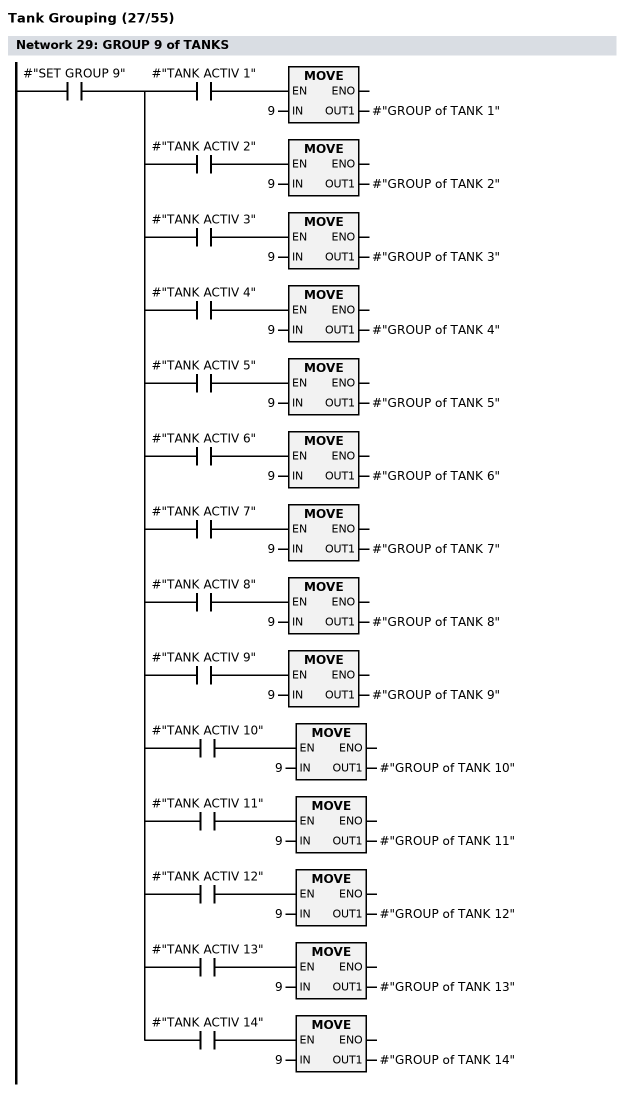
   RUNG wire#powerrail
      Contact( #"SET GROUP 9" )
      wire#w1
      Contact( #"TANK ACTIV 1" )
      Move(in := 9, out1 => #"GROUP of TANK 1")
   END_RUNG
   RUNG wire#w1
      Contact( #"TANK ACTIV 2" )
      Move(in := 9, out1 => #"GROUP of TANK 2")
   END_RUNG
   RUNG wire#w1
      Contact( #"TANK ACTIV 3" )
      Move(in := 9, out1 => #"GROUP of TANK 3")
   END_RUNG
   RUNG wire#w1
      Contact( #"TANK ACTIV 4" )
      Move(in := 9, out1 => #"GROUP of TANK 4")
   END_RUNG
   RUNG wire#w1
      Contact( #"TANK ACTIV 5" )
      Move(in := 9, out1 => #"GROUP of TANK 5")
   END_RUNG
   RUNG wire#w1
      Contact( #"TANK ACTIV 6" )
      Move(in := 9, out1 => #"GROUP of TANK 6")
   END_RUNG
   RUNG wire#w1
      Contact( #"TANK ACTIV 7" )
      Move(in := 9, out1 => #"GROUP of TANK 7")
   END_RUNG
   RUNG wire#w1
      Contact( #"TANK ACTIV 8" )
      Move(in := 9, out1 => #"GROUP of TANK 8")
   END_RUNG
   RUNG wire#w1
      Contact( #"TANK ACTIV 9" )
      Move(in := 9, out1 => #"GROUP of TANK 9")
   END_RUNG
   RUNG wire#w1
      Contact( #"TANK ACTIV 10" )
      Move(in := 9, out1 => #"GROUP of TANK 10")
   END_RUNG
   RUNG wire#w1
      Contact( #"TANK ACTIV 11" )
      Move(in := 9, out1 => #"GROUP of TANK 11")
   END_RUNG
   RUNG wire#w1
      Contact( #"TANK ACTIV 12" )
      Move(in := 9, out1 => #"GROUP of TANK 12")
   END_RUNG
   RUNG wire#w1
      Contact( #"TANK ACTIV 13" )
      Move(in := 9, out1 => #"GROUP of TANK 13")
   END_RUNG
   RUNG wire#w1
      Contact( #"TANK ACTIV 14" )
      Move(in := 9, out1 => #"GROUP of TANK 14")
   END_RUNG
   // the same network as SCL:
   IF #"SET GROUP 9" AND #"TANK ACTIV 1" THEN #"GROUP of TANK 1" := 9; END_IF;
   IF #"SET GROUP 9" AND #"TANK ACTIV 2" THEN #"GROUP of TANK 2" := 9; END_IF;
   IF #"SET GROUP 9" AND #"TANK ACTIV 3" THEN #"GROUP of TANK 3" := 9; END_IF;
   IF #"SET GROUP 9" AND #"TANK ACTIV 4" THEN #"GROUP of TANK 4" := 9; END_IF;
   IF #"SET GROUP 9" AND #"TANK ACTIV 5" THEN #"GROUP of TANK 5" := 9; END_IF;
   IF #"SET GROUP 9" AND #"TANK ACTIV 6" THEN #"GROUP of TANK 6" := 9; END_IF;
   IF #"SET GROUP 9" AND #"TANK ACTIV 7" THEN #"GROUP of TANK 7" := 9; END_IF;
   IF #"SET GROUP 9" AND #"TANK ACTIV 8" THEN #"GROUP of TANK 8" := 9; END_IF;
   IF #"SET GROUP 9" AND #"TANK ACTIV 9" THEN #"GROUP of TANK 9" := 9; END_IF;
   IF #"SET GROUP 9" AND #"TANK ACTIV 10" THEN #"GROUP of TANK 10" := 9; END_IF;
   IF #"SET GROUP 9" AND #"TANK ACTIV 11" THEN #"GROUP of TANK 11" := 9; END_IF;
   IF #"SET GROUP 9" AND #"TANK ACTIV 12" THEN #"GROUP of TANK 12" := 9; END_IF;
   IF #"SET GROUP 9" AND #"TANK ACTIV 13" THEN #"GROUP of TANK 13" := 9; END_IF;
   IF #"SET GROUP 9" AND #"TANK ACTIV 14" THEN #"GROUP of TANK 14" := 9; END_IF;
END_REGION

REGION Network 30: GROUP 10 of TANKS
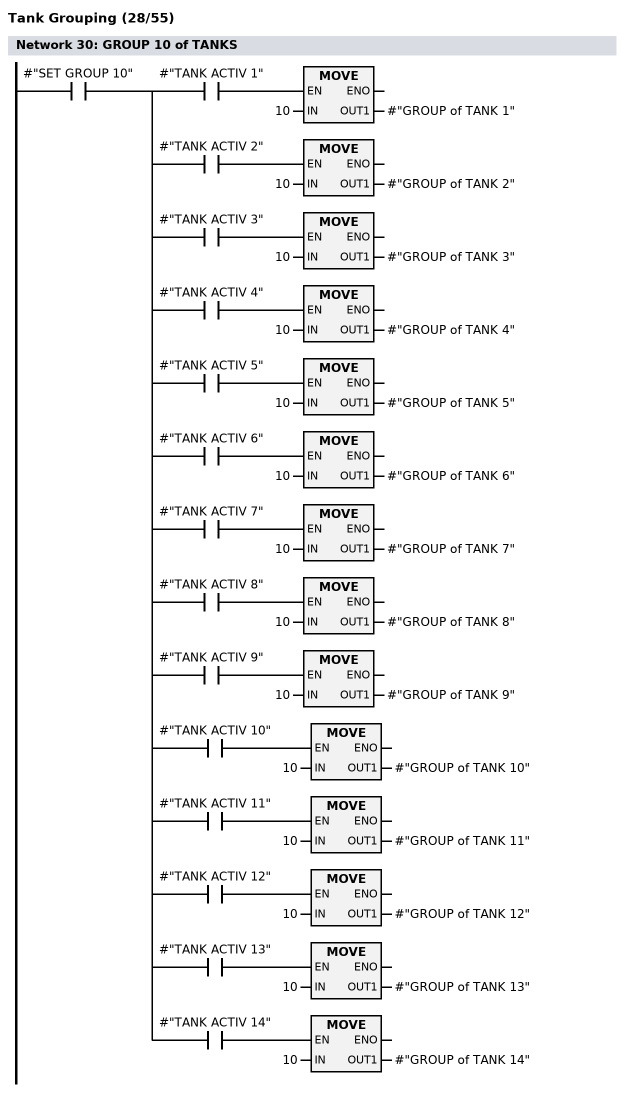
   RUNG wire#powerrail
      Contact( #"SET GROUP 10" )
      wire#w1
      Contact( #"TANK ACTIV 1" )
      Move(in := 10, out1 => #"GROUP of TANK 1")
   END_RUNG
   RUNG wire#w1
      Contact( #"TANK ACTIV 2" )
      Move(in := 10, out1 => #"GROUP of TANK 2")
   END_RUNG
   RUNG wire#w1
      Contact( #"TANK ACTIV 3" )
      Move(in := 10, out1 => #"GROUP of TANK 3")
   END_RUNG
   RUNG wire#w1
      Contact( #"TANK ACTIV 4" )
      Move(in := 10, out1 => #"GROUP of TANK 4")
   END_RUNG
   RUNG wire#w1
      Contact( #"TANK ACTIV 5" )
      Move(in := 10, out1 => #"GROUP of TANK 5")
   END_RUNG
   RUNG wire#w1
      Contact( #"TANK ACTIV 6" )
      Move(in := 10, out1 => #"GROUP of TANK 6")
   END_RUNG
   RUNG wire#w1
      Contact( #"TANK ACTIV 7" )
      Move(in := 10, out1 => #"GROUP of TANK 7")
   END_RUNG
   RUNG wire#w1
      Contact( #"TANK ACTIV 8" )
      Move(in := 10, out1 => #"GROUP of TANK 8")
   END_RUNG
   RUNG wire#w1
      Contact( #"TANK ACTIV 9" )
      Move(in := 10, out1 => #"GROUP of TANK 9")
   END_RUNG
   RUNG wire#w1
      Contact( #"TANK ACTIV 10" )
      Move(in := 10, out1 => #"GROUP of TANK 10")
   END_RUNG
   RUNG wire#w1
      Contact( #"TANK ACTIV 11" )
      Move(in := 10, out1 => #"GROUP of TANK 11")
   END_RUNG
   RUNG wire#w1
      Contact( #"TANK ACTIV 12" )
      Move(in := 10, out1 => #"GROUP of TANK 12")
   END_RUNG
   RUNG wire#w1
      Contact( #"TANK ACTIV 13" )
      Move(in := 10, out1 => #"GROUP of TANK 13")
   END_RUNG
   RUNG wire#w1
      Contact( #"TANK ACTIV 14" )
      Move(in := 10, out1 => #"GROUP of TANK 14")
   END_RUNG
   // the same network as SCL:
   IF #"SET GROUP 10" AND #"TANK ACTIV 1" THEN #"GROUP of TANK 1" := 10; END_IF;
   IF #"SET GROUP 10" AND #"TANK ACTIV 2" THEN #"GROUP of TANK 2" := 10; END_IF;
   IF #"SET GROUP 10" AND #"TANK ACTIV 3" THEN #"GROUP of TANK 3" := 10; END_IF;
   IF #"SET GROUP 10" AND #"TANK ACTIV 4" THEN #"GROUP of TANK 4" := 10; END_IF;
   IF #"SET GROUP 10" AND #"TANK ACTIV 5" THEN #"GROUP of TANK 5" := 10; END_IF;
   IF #"SET GROUP 10" AND #"TANK ACTIV 6" THEN #"GROUP of TANK 6" := 10; END_IF;
   IF #"SET GROUP 10" AND #"TANK ACTIV 7" THEN #"GROUP of TANK 7" := 10; END_IF;
   IF #"SET GROUP 10" AND #"TANK ACTIV 8" THEN #"GROUP of TANK 8" := 10; END_IF;
   IF #"SET GROUP 10" AND #"TANK ACTIV 9" THEN #"GROUP of TANK 9" := 10; END_IF;
   IF #"SET GROUP 10" AND #"TANK ACTIV 10" THEN #"GROUP of TANK 10" := 10; END_IF;
   IF #"SET GROUP 10" AND #"TANK ACTIV 11" THEN #"GROUP of TANK 11" := 10; END_IF;
   IF #"SET GROUP 10" AND #"TANK ACTIV 12" THEN #"GROUP of TANK 12" := 10; END_IF;
   IF #"SET GROUP 10" AND #"TANK ACTIV 13" THEN #"GROUP of TANK 13" := 10; END_IF;
   IF #"SET GROUP 10" AND #"TANK ACTIV 14" THEN #"GROUP of TANK 14" := 10; END_IF;
END_REGION

REGION Network 31: GROUP 11 of TANKS
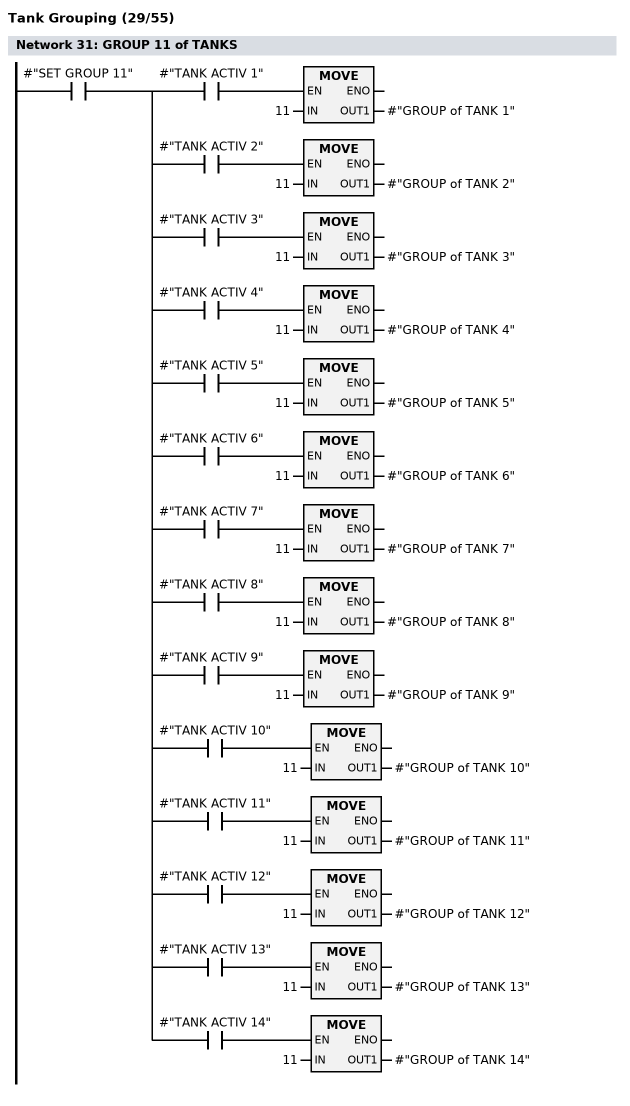
   RUNG wire#powerrail
      Contact( #"SET GROUP 11" )
      wire#w1
      Contact( #"TANK ACTIV 1" )
      Move(in := 11, out1 => #"GROUP of TANK 1")
   END_RUNG
   RUNG wire#w1
      Contact( #"TANK ACTIV 2" )
      Move(in := 11, out1 => #"GROUP of TANK 2")
   END_RUNG
   RUNG wire#w1
      Contact( #"TANK ACTIV 3" )
      Move(in := 11, out1 => #"GROUP of TANK 3")
   END_RUNG
   RUNG wire#w1
      Contact( #"TANK ACTIV 4" )
      Move(in := 11, out1 => #"GROUP of TANK 4")
   END_RUNG
   RUNG wire#w1
      Contact( #"TANK ACTIV 5" )
      Move(in := 11, out1 => #"GROUP of TANK 5")
   END_RUNG
   RUNG wire#w1
      Contact( #"TANK ACTIV 6" )
      Move(in := 11, out1 => #"GROUP of TANK 6")
   END_RUNG
   RUNG wire#w1
      Contact( #"TANK ACTIV 7" )
      Move(in := 11, out1 => #"GROUP of TANK 7")
   END_RUNG
   RUNG wire#w1
      Contact( #"TANK ACTIV 8" )
      Move(in := 11, out1 => #"GROUP of TANK 8")
   END_RUNG
   RUNG wire#w1
      Contact( #"TANK ACTIV 9" )
      Move(in := 11, out1 => #"GROUP of TANK 9")
   END_RUNG
   RUNG wire#w1
      Contact( #"TANK ACTIV 10" )
      Move(in := 11, out1 => #"GROUP of TANK 10")
   END_RUNG
   RUNG wire#w1
      Contact( #"TANK ACTIV 11" )
      Move(in := 11, out1 => #"GROUP of TANK 11")
   END_RUNG
   RUNG wire#w1
      Contact( #"TANK ACTIV 12" )
      Move(in := 11, out1 => #"GROUP of TANK 12")
   END_RUNG
   RUNG wire#w1
      Contact( #"TANK ACTIV 13" )
      Move(in := 11, out1 => #"GROUP of TANK 13")
   END_RUNG
   RUNG wire#w1
      Contact( #"TANK ACTIV 14" )
      Move(in := 11, out1 => #"GROUP of TANK 14")
   END_RUNG
   // the same network as SCL:
   IF #"SET GROUP 11" AND #"TANK ACTIV 1" THEN #"GROUP of TANK 1" := 11; END_IF;
   IF #"SET GROUP 11" AND #"TANK ACTIV 2" THEN #"GROUP of TANK 2" := 11; END_IF;
   IF #"SET GROUP 11" AND #"TANK ACTIV 3" THEN #"GROUP of TANK 3" := 11; END_IF;
   IF #"SET GROUP 11" AND #"TANK ACTIV 4" THEN #"GROUP of TANK 4" := 11; END_IF;
   IF #"SET GROUP 11" AND #"TANK ACTIV 5" THEN #"GROUP of TANK 5" := 11; END_IF;
   IF #"SET GROUP 11" AND #"TANK ACTIV 6" THEN #"GROUP of TANK 6" := 11; END_IF;
   IF #"SET GROUP 11" AND #"TANK ACTIV 7" THEN #"GROUP of TANK 7" := 11; END_IF;
   IF #"SET GROUP 11" AND #"TANK ACTIV 8" THEN #"GROUP of TANK 8" := 11; END_IF;
   IF #"SET GROUP 11" AND #"TANK ACTIV 9" THEN #"GROUP of TANK 9" := 11; END_IF;
   IF #"SET GROUP 11" AND #"TANK ACTIV 10" THEN #"GROUP of TANK 10" := 11; END_IF;
   IF #"SET GROUP 11" AND #"TANK ACTIV 11" THEN #"GROUP of TANK 11" := 11; END_IF;
   IF #"SET GROUP 11" AND #"TANK ACTIV 12" THEN #"GROUP of TANK 12" := 11; END_IF;
   IF #"SET GROUP 11" AND #"TANK ACTIV 13" THEN #"GROUP of TANK 13" := 11; END_IF;
   IF #"SET GROUP 11" AND #"TANK ACTIV 14" THEN #"GROUP of TANK 14" := 11; END_IF;
END_REGION

REGION Network 32: GROUP 12 of TANKS
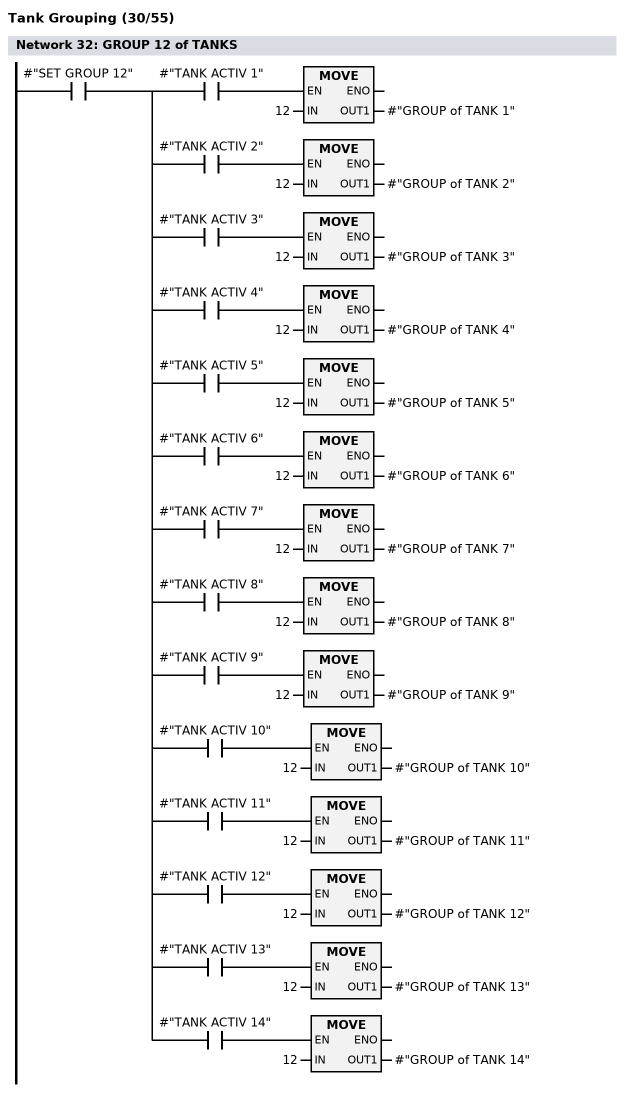
   RUNG wire#powerrail
      Contact( #"SET GROUP 12" )
      wire#w1
      Contact( #"TANK ACTIV 1" )
      Move(in := 12, out1 => #"GROUP of TANK 1")
   END_RUNG
   RUNG wire#w1
      Contact( #"TANK ACTIV 2" )
      Move(in := 12, out1 => #"GROUP of TANK 2")
   END_RUNG
   RUNG wire#w1
      Contact( #"TANK ACTIV 3" )
      Move(in := 12, out1 => #"GROUP of TANK 3")
   END_RUNG
   RUNG wire#w1
      Contact( #"TANK ACTIV 4" )
      Move(in := 12, out1 => #"GROUP of TANK 4")
   END_RUNG
   RUNG wire#w1
      Contact( #"TANK ACTIV 5" )
      Move(in := 12, out1 => #"GROUP of TANK 5")
   END_RUNG
   RUNG wire#w1
      Contact( #"TANK ACTIV 6" )
      Move(in := 12, out1 => #"GROUP of TANK 6")
   END_RUNG
   RUNG wire#w1
      Contact( #"TANK ACTIV 7" )
      Move(in := 12, out1 => #"GROUP of TANK 7")
   END_RUNG
   RUNG wire#w1
      Contact( #"TANK ACTIV 8" )
      Move(in := 12, out1 => #"GROUP of TANK 8")
   END_RUNG
   RUNG wire#w1
      Contact( #"TANK ACTIV 9" )
      Move(in := 12, out1 => #"GROUP of TANK 9")
   END_RUNG
   RUNG wire#w1
      Contact( #"TANK ACTIV 10" )
      Move(in := 12, out1 => #"GROUP of TANK 10")
   END_RUNG
   RUNG wire#w1
      Contact( #"TANK ACTIV 11" )
      Move(in := 12, out1 => #"GROUP of TANK 11")
   END_RUNG
   RUNG wire#w1
      Contact( #"TANK ACTIV 12" )
      Move(in := 12, out1 => #"GROUP of TANK 12")
   END_RUNG
   RUNG wire#w1
      Contact( #"TANK ACTIV 13" )
      Move(in := 12, out1 => #"GROUP of TANK 13")
   END_RUNG
   RUNG wire#w1
      Contact( #"TANK ACTIV 14" )
      Move(in := 12, out1 => #"GROUP of TANK 14")
   END_RUNG
   // the same network as SCL:
   IF #"SET GROUP 12" AND #"TANK ACTIV 1" THEN #"GROUP of TANK 1" := 12; END_IF;
   IF #"SET GROUP 12" AND #"TANK ACTIV 2" THEN #"GROUP of TANK 2" := 12; END_IF;
   IF #"SET GROUP 12" AND #"TANK ACTIV 3" THEN #"GROUP of TANK 3" := 12; END_IF;
   IF #"SET GROUP 12" AND #"TANK ACTIV 4" THEN #"GROUP of TANK 4" := 12; END_IF;
   IF #"SET GROUP 12" AND #"TANK ACTIV 5" THEN #"GROUP of TANK 5" := 12; END_IF;
   IF #"SET GROUP 12" AND #"TANK ACTIV 6" THEN #"GROUP of TANK 6" := 12; END_IF;
   IF #"SET GROUP 12" AND #"TANK ACTIV 7" THEN #"GROUP of TANK 7" := 12; END_IF;
   IF #"SET GROUP 12" AND #"TANK ACTIV 8" THEN #"GROUP of TANK 8" := 12; END_IF;
   IF #"SET GROUP 12" AND #"TANK ACTIV 9" THEN #"GROUP of TANK 9" := 12; END_IF;
   IF #"SET GROUP 12" AND #"TANK ACTIV 10" THEN #"GROUP of TANK 10" := 12; END_IF;
   IF #"SET GROUP 12" AND #"TANK ACTIV 11" THEN #"GROUP of TANK 11" := 12; END_IF;
   IF #"SET GROUP 12" AND #"TANK ACTIV 12" THEN #"GROUP of TANK 12" := 12; END_IF;
   IF #"SET GROUP 12" AND #"TANK ACTIV 13" THEN #"GROUP of TANK 13" := 12; END_IF;
   IF #"SET GROUP 12" AND #"TANK ACTIV 14" THEN #"GROUP of TANK 14" := 12; END_IF;
END_REGION

REGION Network 33: GROUP 13 of TANKS
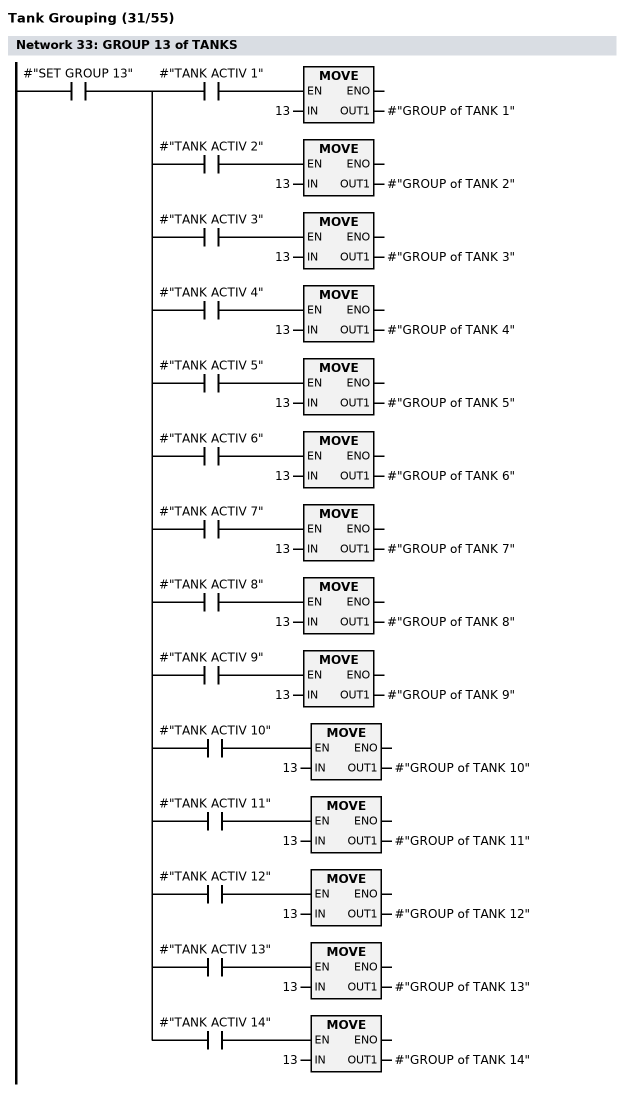
   RUNG wire#powerrail
      Contact( #"SET GROUP 13" )
      wire#w1
      Contact( #"TANK ACTIV 1" )
      Move(in := 13, out1 => #"GROUP of TANK 1")
   END_RUNG
   RUNG wire#w1
      Contact( #"TANK ACTIV 2" )
      Move(in := 13, out1 => #"GROUP of TANK 2")
   END_RUNG
   RUNG wire#w1
      Contact( #"TANK ACTIV 3" )
      Move(in := 13, out1 => #"GROUP of TANK 3")
   END_RUNG
   RUNG wire#w1
      Contact( #"TANK ACTIV 4" )
      Move(in := 13, out1 => #"GROUP of TANK 4")
   END_RUNG
   RUNG wire#w1
      Contact( #"TANK ACTIV 5" )
      Move(in := 13, out1 => #"GROUP of TANK 5")
   END_RUNG
   RUNG wire#w1
      Contact( #"TANK ACTIV 6" )
      Move(in := 13, out1 => #"GROUP of TANK 6")
   END_RUNG
   RUNG wire#w1
      Contact( #"TANK ACTIV 7" )
      Move(in := 13, out1 => #"GROUP of TANK 7")
   END_RUNG
   RUNG wire#w1
      Contact( #"TANK ACTIV 8" )
      Move(in := 13, out1 => #"GROUP of TANK 8")
   END_RUNG
   RUNG wire#w1
      Contact( #"TANK ACTIV 9" )
      Move(in := 13, out1 => #"GROUP of TANK 9")
   END_RUNG
   RUNG wire#w1
      Contact( #"TANK ACTIV 10" )
      Move(in := 13, out1 => #"GROUP of TANK 10")
   END_RUNG
   RUNG wire#w1
      Contact( #"TANK ACTIV 11" )
      Move(in := 13, out1 => #"GROUP of TANK 11")
   END_RUNG
   RUNG wire#w1
      Contact( #"TANK ACTIV 12" )
      Move(in := 13, out1 => #"GROUP of TANK 12")
   END_RUNG
   RUNG wire#w1
      Contact( #"TANK ACTIV 13" )
      Move(in := 13, out1 => #"GROUP of TANK 13")
   END_RUNG
   RUNG wire#w1
      Contact( #"TANK ACTIV 14" )
      Move(in := 13, out1 => #"GROUP of TANK 14")
   END_RUNG
   // the same network as SCL:
   IF #"SET GROUP 13" AND #"TANK ACTIV 1" THEN #"GROUP of TANK 1" := 13; END_IF;
   IF #"SET GROUP 13" AND #"TANK ACTIV 2" THEN #"GROUP of TANK 2" := 13; END_IF;
   IF #"SET GROUP 13" AND #"TANK ACTIV 3" THEN #"GROUP of TANK 3" := 13; END_IF;
   IF #"SET GROUP 13" AND #"TANK ACTIV 4" THEN #"GROUP of TANK 4" := 13; END_IF;
   IF #"SET GROUP 13" AND #"TANK ACTIV 5" THEN #"GROUP of TANK 5" := 13; END_IF;
   IF #"SET GROUP 13" AND #"TANK ACTIV 6" THEN #"GROUP of TANK 6" := 13; END_IF;
   IF #"SET GROUP 13" AND #"TANK ACTIV 7" THEN #"GROUP of TANK 7" := 13; END_IF;
   IF #"SET GROUP 13" AND #"TANK ACTIV 8" THEN #"GROUP of TANK 8" := 13; END_IF;
   IF #"SET GROUP 13" AND #"TANK ACTIV 9" THEN #"GROUP of TANK 9" := 13; END_IF;
   IF #"SET GROUP 13" AND #"TANK ACTIV 10" THEN #"GROUP of TANK 10" := 13; END_IF;
   IF #"SET GROUP 13" AND #"TANK ACTIV 11" THEN #"GROUP of TANK 11" := 13; END_IF;
   IF #"SET GROUP 13" AND #"TANK ACTIV 12" THEN #"GROUP of TANK 12" := 13; END_IF;
   IF #"SET GROUP 13" AND #"TANK ACTIV 13" THEN #"GROUP of TANK 13" := 13; END_IF;
   IF #"SET GROUP 13" AND #"TANK ACTIV 14" THEN #"GROUP of TANK 14" := 13; END_IF;
END_REGION

REGION Network 34: GROUP 14 of TANKS
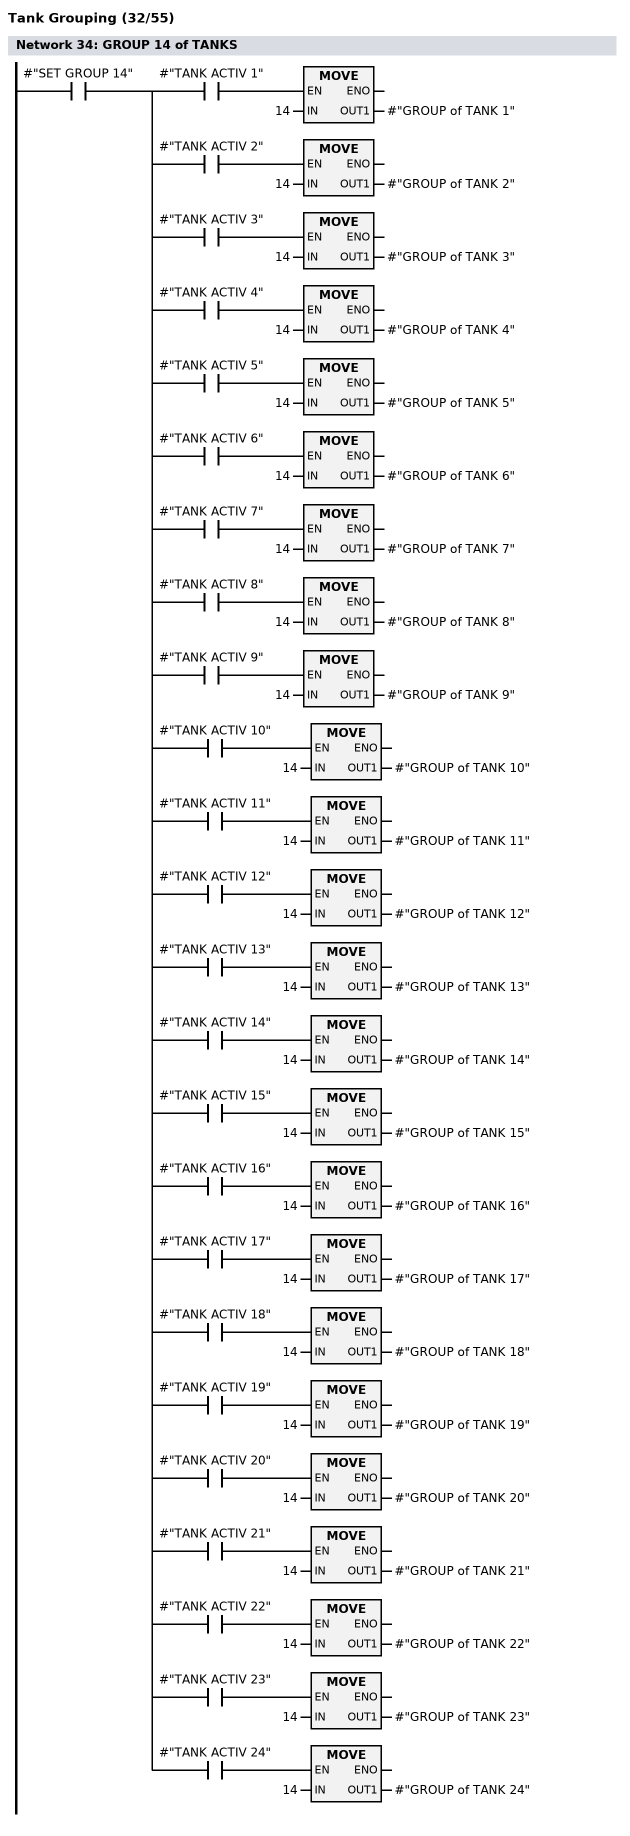
   RUNG wire#powerrail
      Contact( #"SET GROUP 14" )
      wire#w1
      Contact( #"TANK ACTIV 1" )
      Move(in := 14, out1 => #"GROUP of TANK 1")
   END_RUNG
   RUNG wire#w1
      Contact( #"TANK ACTIV 2" )
      Move(in := 14, out1 => #"GROUP of TANK 2")
   END_RUNG
   RUNG wire#w1
      Contact( #"TANK ACTIV 3" )
      Move(in := 14, out1 => #"GROUP of TANK 3")
   END_RUNG
   RUNG wire#w1
      Contact( #"TANK ACTIV 4" )
      Move(in := 14, out1 => #"GROUP of TANK 4")
   END_RUNG
   RUNG wire#w1
      Contact( #"TANK ACTIV 5" )
      Move(in := 14, out1 => #"GROUP of TANK 5")
   END_RUNG
   RUNG wire#w1
      Contact( #"TANK ACTIV 6" )
      Move(in := 14, out1 => #"GROUP of TANK 6")
   END_RUNG
   RUNG wire#w1
      Contact( #"TANK ACTIV 7" )
      Move(in := 14, out1 => #"GROUP of TANK 7")
   END_RUNG
   RUNG wire#w1
      Contact( #"TANK ACTIV 8" )
      Move(in := 14, out1 => #"GROUP of TANK 8")
   END_RUNG
   RUNG wire#w1
      Contact( #"TANK ACTIV 9" )
      Move(in := 14, out1 => #"GROUP of TANK 9")
   END_RUNG
   RUNG wire#w1
      Contact( #"TANK ACTIV 10" )
      Move(in := 14, out1 => #"GROUP of TANK 10")
   END_RUNG
   RUNG wire#w1
      Contact( #"TANK ACTIV 11" )
      Move(in := 14, out1 => #"GROUP of TANK 11")
   END_RUNG
   RUNG wire#w1
      Contact( #"TANK ACTIV 12" )
      Move(in := 14, out1 => #"GROUP of TANK 12")
   END_RUNG
   RUNG wire#w1
      Contact( #"TANK ACTIV 13" )
      Move(in := 14, out1 => #"GROUP of TANK 13")
   END_RUNG
   RUNG wire#w1
      Contact( #"TANK ACTIV 14" )
      Move(in := 14, out1 => #"GROUP of TANK 14")
   END_RUNG
   RUNG wire#w1
      Contact( #"TANK ACTIV 15" )
      Move(in := 14, out1 => #"GROUP of TANK 15")
   END_RUNG
   RUNG wire#w1
      Contact( #"TANK ACTIV 16" )
      Move(in := 14, out1 => #"GROUP of TANK 16")
   END_RUNG
   RUNG wire#w1
      Contact( #"TANK ACTIV 17" )
      Move(in := 14, out1 => #"GROUP of TANK 17")
   END_RUNG
   RUNG wire#w1
      Contact( #"TANK ACTIV 18" )
      Move(in := 14, out1 => #"GROUP of TANK 18")
   END_RUNG
   RUNG wire#w1
      Contact( #"TANK ACTIV 19" )
      Move(in := 14, out1 => #"GROUP of TANK 19")
   END_RUNG
   RUNG wire#w1
      Contact( #"TANK ACTIV 20" )
      Move(in := 14, out1 => #"GROUP of TANK 20")
   END_RUNG
   RUNG wire#w1
      Contact( #"TANK ACTIV 21" )
      Move(in := 14, out1 => #"GROUP of TANK 21")
   END_RUNG
   RUNG wire#w1
      Contact( #"TANK ACTIV 22" )
      Move(in := 14, out1 => #"GROUP of TANK 22")
   END_RUNG
   RUNG wire#w1
      Contact( #"TANK ACTIV 23" )
      Move(in := 14, out1 => #"GROUP of TANK 23")
   END_RUNG
   RUNG wire#w1
      Contact( #"TANK ACTIV 24" )
      Move(in := 14, out1 => #"GROUP of TANK 24")
   END_RUNG
   // the same network as SCL:
   IF #"SET GROUP 14" AND #"TANK ACTIV 1" THEN #"GROUP of TANK 1" := 14; END_IF;
   IF #"SET GROUP 14" AND #"TANK ACTIV 2" THEN #"GROUP of TANK 2" := 14; END_IF;
   IF #"SET GROUP 14" AND #"TANK ACTIV 3" THEN #"GROUP of TANK 3" := 14; END_IF;
   IF #"SET GROUP 14" AND #"TANK ACTIV 4" THEN #"GROUP of TANK 4" := 14; END_IF;
   IF #"SET GROUP 14" AND #"TANK ACTIV 5" THEN #"GROUP of TANK 5" := 14; END_IF;
   IF #"SET GROUP 14" AND #"TANK ACTIV 6" THEN #"GROUP of TANK 6" := 14; END_IF;
   IF #"SET GROUP 14" AND #"TANK ACTIV 7" THEN #"GROUP of TANK 7" := 14; END_IF;
   IF #"SET GROUP 14" AND #"TANK ACTIV 8" THEN #"GROUP of TANK 8" := 14; END_IF;
   IF #"SET GROUP 14" AND #"TANK ACTIV 9" THEN #"GROUP of TANK 9" := 14; END_IF;
   IF #"SET GROUP 14" AND #"TANK ACTIV 10" THEN #"GROUP of TANK 10" := 14; END_IF;
   IF #"SET GROUP 14" AND #"TANK ACTIV 11" THEN #"GROUP of TANK 11" := 14; END_IF;
   IF #"SET GROUP 14" AND #"TANK ACTIV 12" THEN #"GROUP of TANK 12" := 14; END_IF;
   IF #"SET GROUP 14" AND #"TANK ACTIV 13" THEN #"GROUP of TANK 13" := 14; END_IF;
   IF #"SET GROUP 14" AND #"TANK ACTIV 14" THEN #"GROUP of TANK 14" := 14; END_IF;
   IF #"SET GROUP 14" AND #"TANK ACTIV 15" THEN #"GROUP of TANK 15" := 14; END_IF;
   IF #"SET GROUP 14" AND #"TANK ACTIV 16" THEN #"GROUP of TANK 16" := 14; END_IF;
   IF #"SET GROUP 14" AND #"TANK ACTIV 17" THEN #"GROUP of TANK 17" := 14; END_IF;
   IF #"SET GROUP 14" AND #"TANK ACTIV 18" THEN #"GROUP of TANK 18" := 14; END_IF;
   IF #"SET GROUP 14" AND #"TANK ACTIV 19" THEN #"GROUP of TANK 19" := 14; END_IF;
   IF #"SET GROUP 14" AND #"TANK ACTIV 20" THEN #"GROUP of TANK 20" := 14; END_IF;
   IF #"SET GROUP 14" AND #"TANK ACTIV 21" THEN #"GROUP of TANK 21" := 14; END_IF;
   IF #"SET GROUP 14" AND #"TANK ACTIV 22" THEN #"GROUP of TANK 22" := 14; END_IF;
   IF #"SET GROUP 14" AND #"TANK ACTIV 23" THEN #"GROUP of TANK 23" := 14; END_IF;
   IF #"SET GROUP 14" AND #"TANK ACTIV 24" THEN #"GROUP of TANK 24" := 14; END_IF;
END_REGION

REGION Network 35: RESET & MEMORY of TANKS
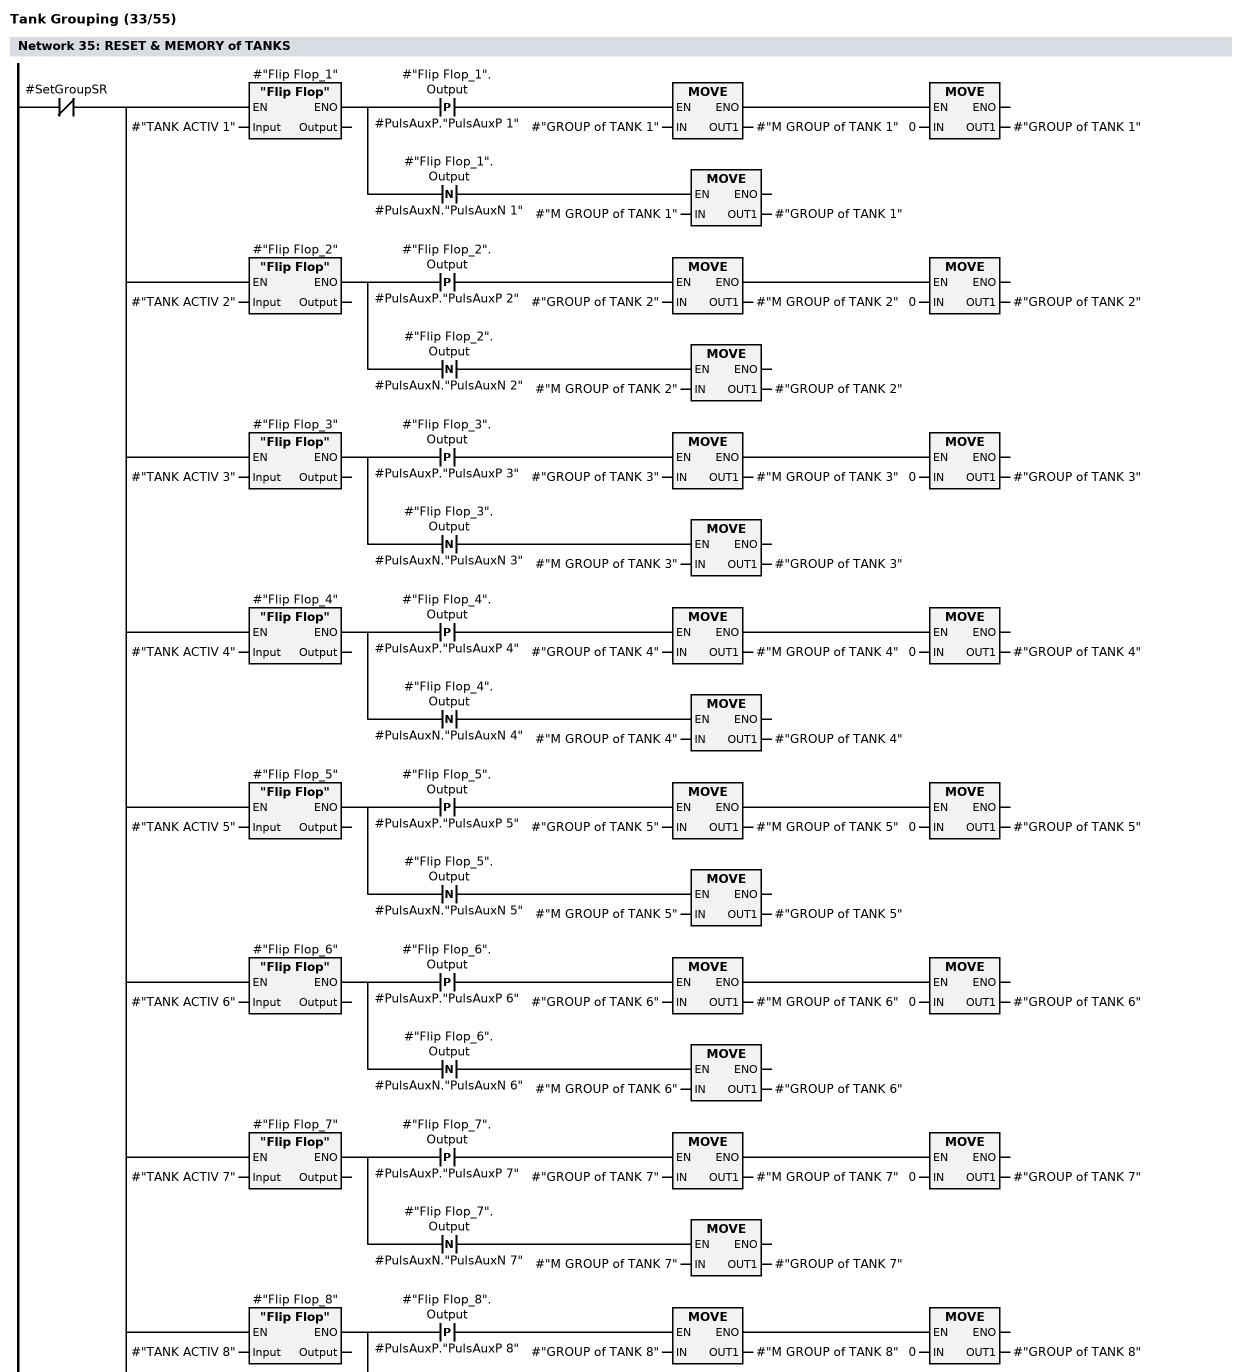